// TIA Portal project "TestEssProtoFreia" (V13) (continued)
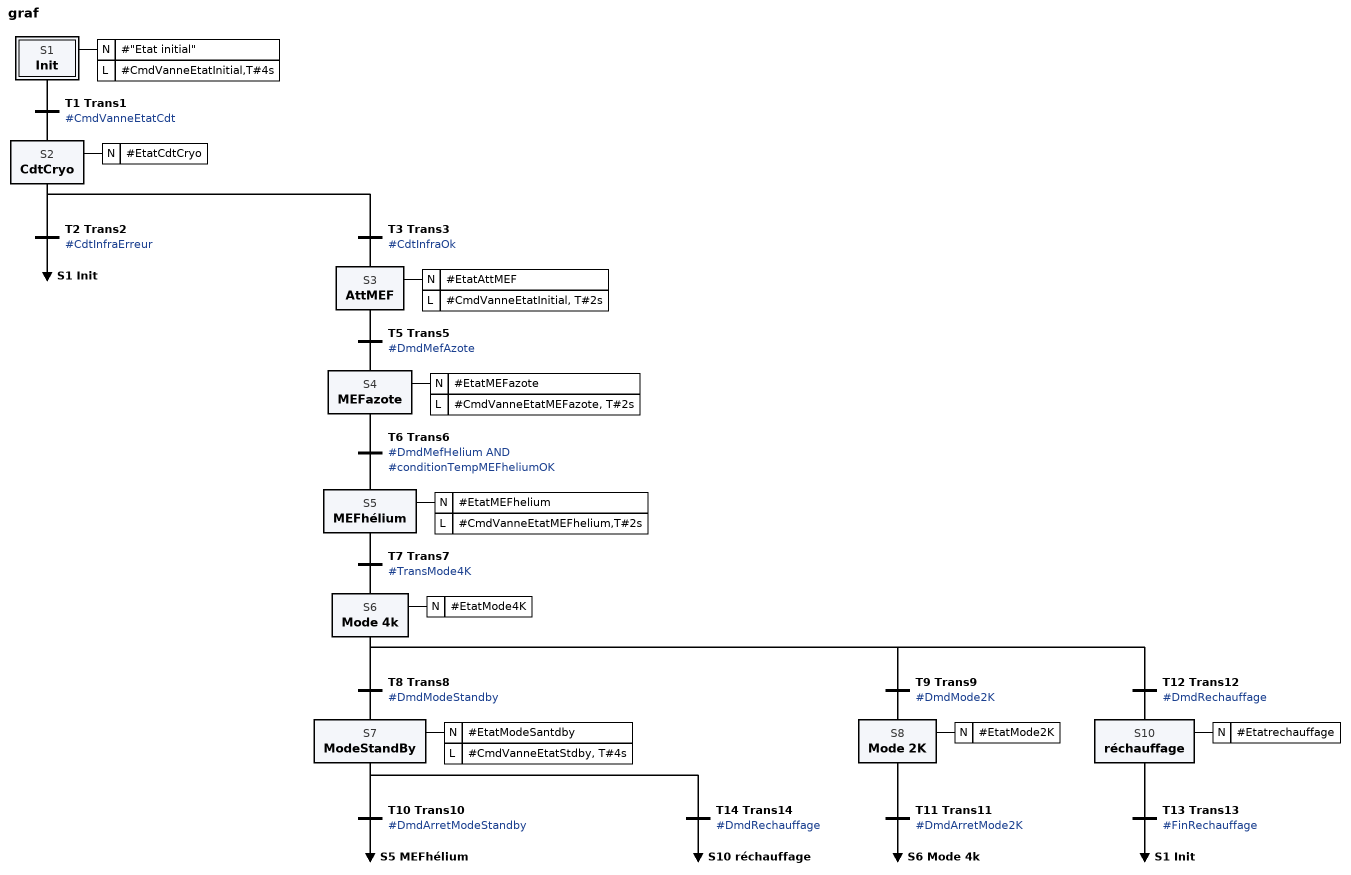
   // sequencer 1
   INITIAL_STEP Init:   // S1
              N    #"Etat initial"
              L    #CmdVanneEtatInitial,T#4s
   END_STEP
   TRANSITION Trans1 FROM Init TO CdtCryo   // T1
      := #CmdVanneEtatCdt;
   END_TRANSITION
   STEP CdtCryo:   // S2
      supervision V := NOT #VanneEnPositionCdt;
      // Version 1: demander manuellement à l automate infra de faire le cdt et confirmer manuellement ( ou pas ) le conditionnement trans3 ( ou trans 2 ) [ajouter boutton cdtinfraok et cdtinfra erreur]
              N    #EtatCdtCryo
   END_STEP
   TRANSITION Trans2 FROM CdtCryo TO Init   // T2, jump
      := #CdtInfraErreur;
   END_TRANSITION
   TRANSITION Trans3 FROM CdtCryo TO AttMEF   // T3
      := #CdtInfraOk;
   END_TRANSITION
   STEP AttMEF:   // S3
      supervision V := NOT #AutorizationMefAzote;
              N    #EtatAttMEF
              L    #CmdVanneEtatInitial, T#2s
   END_STEP
   TRANSITION Trans5 FROM AttMEF TO MEFazote   // T5
      := #DmdMefAzote;
   END_TRANSITION
   STEP MEFazote:   // S4
              N    #EtatMEFazote
              L    #CmdVanneEtatMEFazote, T#2s
   END_STEP
   TRANSITION Trans6 FROM MEFazote TO MEFhélium   // T6
      := #DmdMefHelium AND #conditionTempMEFheliumOK;
   END_TRANSITION
   STEP MEFhélium:   // S5
              N    #EtatMEFhelium
              L    #CmdVanneEtatMEFhelium,T#2s
   END_STEP
   TRANSITION Trans7 FROM MEFhélium TO "Mode 4k"   // T7
      := #TransMode4K;
   END_TRANSITION
   STEP "Mode 4k":   // S6
              N    #EtatMode4K
   END_STEP
   TRANSITION Trans8 FROM "Mode 4k" TO ModeStandBy   // T8
      := #DmdModeStandby;
   END_TRANSITION
   TRANSITION Trans9 FROM "Mode 4k" TO "Mode 2K"   // T9
      := #DmdMode2K;
   END_TRANSITION
   TRANSITION Trans12 FROM "Mode 4k" TO réchauffage   // T12
      := #DmdRechauffage;
   END_TRANSITION
   STEP ModeStandBy:   // S7
              N    #EtatModeSantdby
              L    #CmdVanneEtatStdby, T#4s
   END_STEP
   TRANSITION Trans10 FROM ModeStandBy TO MEFhélium   // T10, jump
      := #DmdArretModeStandby;
   END_TRANSITION
   TRANSITION Trans14 FROM ModeStandBy TO réchauffage   // T14, jump
      := #DmdRechauffage;
   END_TRANSITION
   STEP "Mode 2K":   // S8
              N    #EtatMode2K
   END_STEP
   TRANSITION Trans11 FROM "Mode 2K" TO "Mode 4k"   // T11, jump
      := #DmdArretMode2K;
   END_TRANSITION
   STEP réchauffage:   // S10
              N    #Etatrechauffage
   END_STEP
   TRANSITION Trans13 FROM réchauffage TO Init   // T13, jump
      := #FinRechauffage;
   END_TRANSITION
END_FUNCTION_BLOCK

FUNCTION "commande vanne" : Void   // FC1, LAD
{ S7_Optimized_Access := 'FALSE' }
VERSION : 0.1
   VAR_TEMP   // added for the SCL form of the ladder/FBD networks
      _w1 : Bool;
   END_VAR
BEGIN

REGION Network 1: CV01
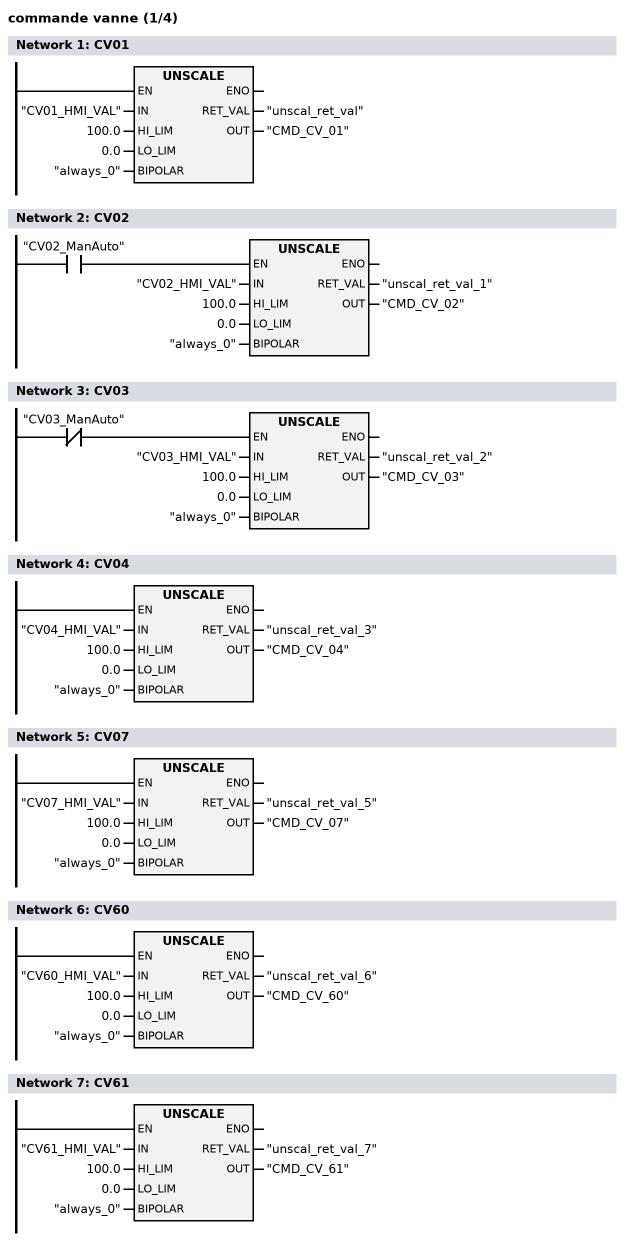
   "unscal_ret_val" := UNSCALE(IN := "CV01_HMI_VAL",
                           HI_LIM := 100.0,
                           LO_LIM := 0.0,
                           BIPOLAR := "always_0",
                           OUT => "CMD_CV_01");
END_REGION

REGION Network 2: CV02
   IF "CV02_ManAuto" THEN
       "unscal_ret_val_1" := UNSCALE(IN := "CV02_HMI_VAL",
                               HI_LIM := 100.0,
                               LO_LIM := 0.0,
                               BIPOLAR := "always_0",
                               OUT => "CMD_CV_02");
   END_IF;
END_REGION

REGION Network 3: CV03
   IF NOT "CV03_ManAuto" THEN
       "unscal_ret_val_2" := UNSCALE(IN := "CV03_HMI_VAL",
                               HI_LIM := 100.0,
                               LO_LIM := 0.0,
                               BIPOLAR := "always_0",
                               OUT => "CMD_CV_03");
   END_IF;
END_REGION

REGION Network 4: CV04
   "unscal_ret_val_3" := UNSCALE(IN := "CV04_HMI_VAL",
                           HI_LIM := 100.0,
                           LO_LIM := 0.0,
                           BIPOLAR := "always_0",
                           OUT => "CMD_CV_04");
END_REGION

REGION Network 5: CV07
   "unscal_ret_val_5" := UNSCALE(IN := "CV07_HMI_VAL",
                           HI_LIM := 100.0,
                           LO_LIM := 0.0,
                           BIPOLAR := "always_0",
                           OUT => "CMD_CV_07");
END_REGION

REGION Network 6: CV60
   "unscal_ret_val_6" := UNSCALE(IN := "CV60_HMI_VAL",
                           HI_LIM := 100.0,
                           LO_LIM := 0.0,
                           BIPOLAR := "always_0",
                           OUT => "CMD_CV_60");
END_REGION

REGION Network 7: CV61
   "unscal_ret_val_7" := UNSCALE(IN := "CV61_HMI_VAL",
                           HI_LIM := 100.0,
                           LO_LIM := 0.0,
                           BIPOLAR := "always_0",
                           OUT => "CMD_CV_61");
END_REGION

REGION Network 8: FT11 (CV11)
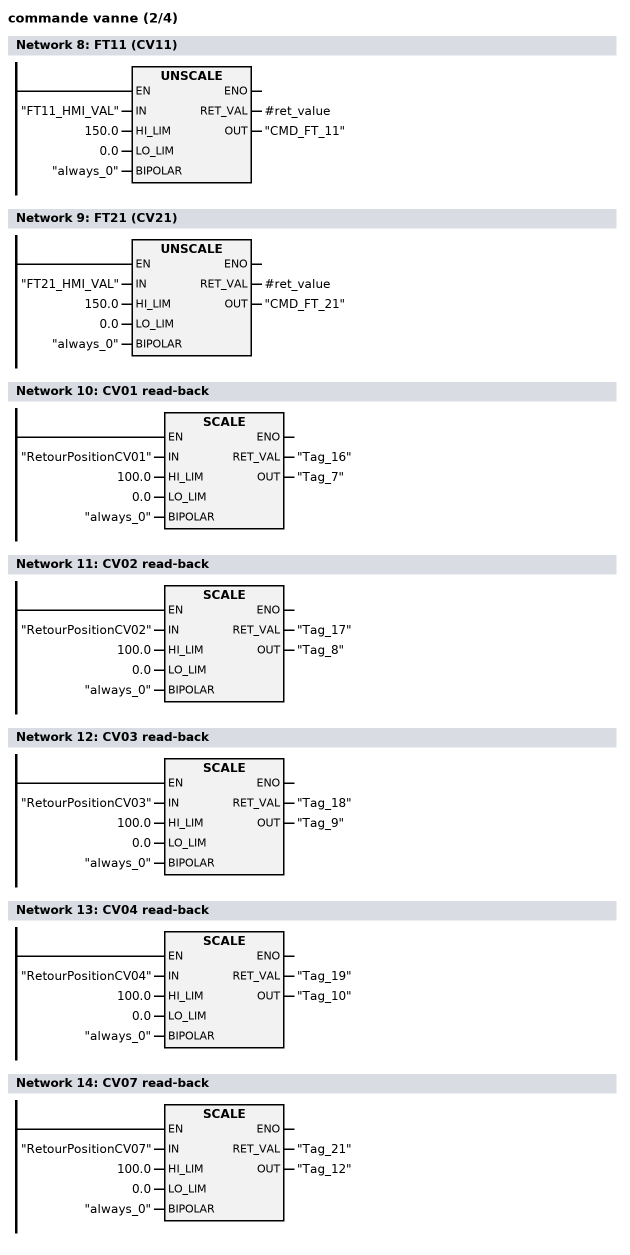
   #ret_value := UNSCALE(IN := "FT11_HMI_VAL",
                         HI_LIM := 150.0,
                         LO_LIM := 0.0,
                         BIPOLAR := "always_0",
                         OUT => "CMD_FT_11");
END_REGION

REGION Network 9: FT21 (CV21)
   #ret_value := UNSCALE(IN := "FT21_HMI_VAL",
                         HI_LIM := 150.0,
                         LO_LIM := 0.0,
                         BIPOLAR := "always_0",
                         OUT => "CMD_FT_21");
END_REGION

REGION Network 10: CV01 read-back
   "Tag_16" := SCALE(IN := "RetourPositionCV01",
                     HI_LIM := 100.0,
                     LO_LIM := 0.0,
                     BIPOLAR := "always_0",
                     OUT => "Tag_7");
END_REGION

REGION Network 11: CV02 read-back
   "Tag_17" := SCALE(IN := "RetourPositionCV02",
                     HI_LIM := 100.0,
                     LO_LIM := 0.0,
                     BIPOLAR := "always_0",
                     OUT => "Tag_8");
END_REGION

REGION Network 12: CV03 read-back
   "Tag_18" := SCALE(IN := "RetourPositionCV03",
                     HI_LIM := 100.0,
                     LO_LIM := 0.0,
                     BIPOLAR := "always_0",
                     OUT => "Tag_9");
END_REGION

REGION Network 13: CV04 read-back
   "Tag_19" := SCALE(IN := "RetourPositionCV04",
                     HI_LIM := 100.0,
                     LO_LIM := 0.0,
                     BIPOLAR := "always_0",
                     OUT => "Tag_10");
END_REGION

REGION Network 14: CV07 read-back
   "Tag_21" := SCALE(IN := "RetourPositionCV07",
                     HI_LIM := 100.0,
                     LO_LIM := 0.0,
                     BIPOLAR := "always_0",
                     OUT => "Tag_12");
END_REGION

REGION Network 15: CV60 read-back
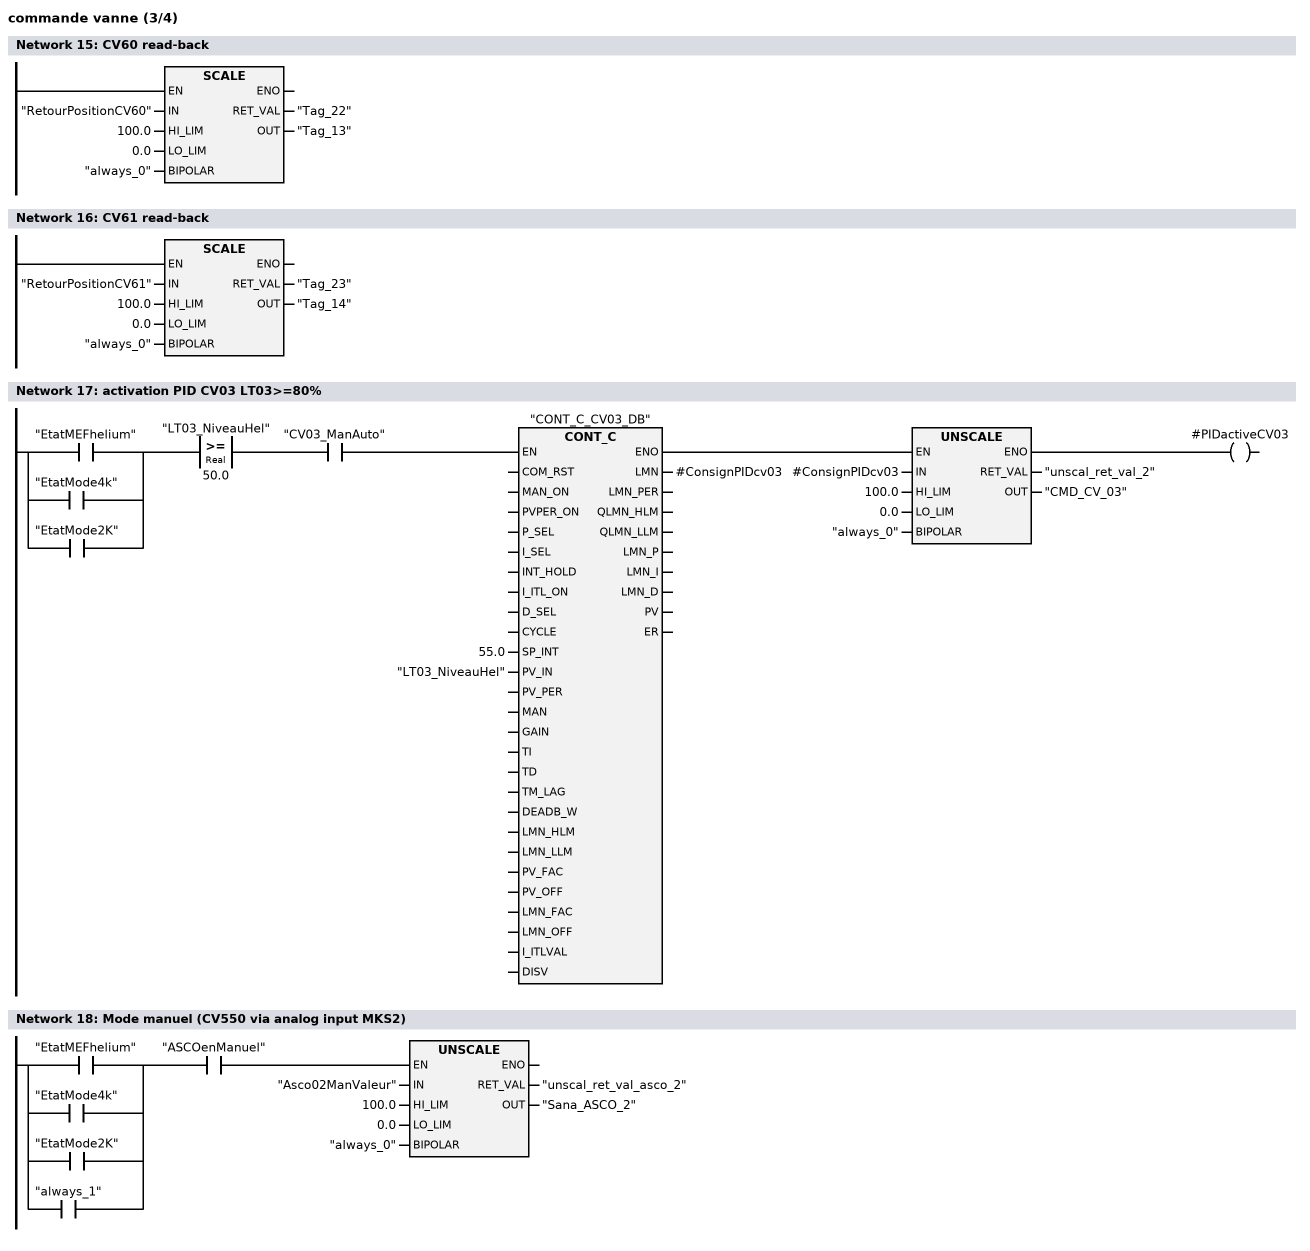
   "Tag_22" := SCALE(IN := "RetourPositionCV60",
                     HI_LIM := 100.0,
                     LO_LIM := 0.0,
                     BIPOLAR := "always_0",
                     OUT => "Tag_13");
END_REGION

REGION Network 16: CV61 read-back
   "Tag_23" := SCALE(IN := "RetourPositionCV61",
                     HI_LIM := 100.0,
                     LO_LIM := 0.0,
                     BIPOLAR := "always_0",
                     OUT => "Tag_14");
END_REGION

REGION Network 17: activation PID CV03 LT03>=80%
   // ENO of a box is taken as its EN; it also drops when the box reports an error
   #_w1 := ("EtatMEFhelium" OR "EtatMode4k" OR "EtatMode2K") AND ("LT03_NiveauHel" >= 50.0) AND "CV03_ManAuto";
   IF #_w1 THEN
       "CONT_C_CV03_DB"(SP_INT := 55.0, PV_IN := "LT03_NiveauHel", LMN => #ConsignPIDcv03);   // CONT_C
       "unscal_ret_val_2" := UNSCALE(IN := #ConsignPIDcv03,
                               HI_LIM := 100.0,
                               LO_LIM := 0.0,
                               BIPOLAR := "always_0",
                               OUT => "CMD_CV_03");
   END_IF;
   #PIDactiveCV03 := #_w1;
END_REGION

REGION Network 18: Mode manuel (CV550 via analog input MKS2)
   IF ("EtatMEFhelium" OR "EtatMode4k" OR "EtatMode2K" OR "always_1") AND "ASCOenManuel" THEN
       "unscal_ret_val_asco_2" := UNSCALE(IN := "Asco02ManValeur",
                               HI_LIM := 100.0,
                               LO_LIM := 0.0,
                               BIPOLAR := "always_0",
                               OUT => "Sana_ASCO_2");
   END_IF;
END_REGION

REGION Network 19: ASCO2 read-back (CV550 read-back via analog output from MKS2)
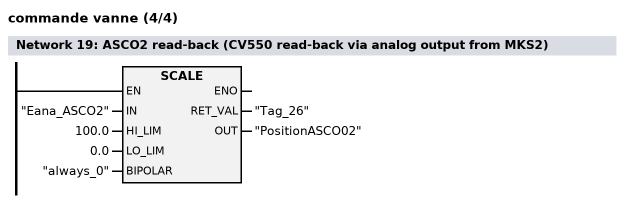
   "Tag_26" := SCALE(IN := "Eana_ASCO2",
                     HI_LIM := 100.0,
                     LO_LIM := 0.0,
                     BIPOLAR := "always_0",
                     OUT => "PositionASCO02");
END_REGION
END_FUNCTION

FUNCTION "NIveau Helium&Pression&vide" : Void   // FC2, STL
{ S7_Optimized_Access := 'FALSE' }
VERSION : 0.1
BEGIN

REGION Network 1: scale niveau helieum LT03
         A     "always_1";
         =     #tmpb;
         BLD   103;
         CALL  "FC10=SCALE"
         ( INPUT       := "Eana_NiveauH_LT03",
           VAL_MAXI    := 74.0,
           VAL_MINI    := 0.0,
           ET_MAX      := 27648,
           ET_MIN      := 0,
           Type_Entree := 0,
           PV_SEUILH   := 100.0,
           PV_SEUILB   := 0.0,
           ACQ         := #tmpb,
           ANIM        := "LT03_TypeDef",
           PV_HIGH     := "LT03_ValMax",
           PV_LOW      := "LT03_ValMin",
           PV          := "LT03_NiveauHel",
           ALM_HIGH    := "LT03_DepHaut",
           ALM_LOW     := "LT03_DepBas",
           ALM_SENSOR  := "LT03_DefSond"
         );
         NOP   0;
END_REGION

REGION Network 2: Copy LT03 to Epics
         L     "LT03_NiveauHel";
         T     "PLC_to_Epics".LT03.Level;
         L     "LT03_TypeDef";
         T     "PLC_to_Epics".LT03.Visu;
         A     "LT03_DefSond";
         =     "PLC_to_Epics".LT03.SensorFlt;
         A     "LT03_DepHaut";
         =     "PLC_to_Epics".LT03.OverRange;
         A     "LT03_DepBas";
         =     "PLC_to_Epics".LT03.UnderRange;
END_REGION

REGION Network 3: scale niveau helieum LT01
         A     "always_1";
         =     #tmpb;
         BLD   103;
         CALL  "FC10=SCALE"
         ( INPUT       := "Eana_NiveauH_LT01",
           VAL_MAXI    := 68.0,
           VAL_MINI    := 0.0,
           ET_MAX      := 27648,
           ET_MIN      := 0,
           Type_Entree := 0,
           PV_SEUILH   := 100.0,
           PV_SEUILB   := 0.0,
           ACQ         := #tmpb,
           ANIM        := "LT01_TypeDef",
           PV_HIGH     := "LT01_ValMax",
           PV_LOW      := "LT01_ValMin",
           PV          := "LT01_NiveauHel",
           ALM_HIGH    := "LT01_DepHaut",
           ALM_LOW     := "LT01_DepBas",
           ALM_SENSOR  := "LT01_DefSond"
         );
         NOP   0;
END_REGION

REGION Network 4: Copy LT01 to Epics
         L     "LT01_NiveauHel";
         T     "PLC_to_Epics".LT01.Level;
         L     "LT01_TypeDef";
         T     "PLC_to_Epics".LT01.Visu;
         A     "LT01_DefSond";
         =     "PLC_to_Epics".LT01.SensorFlt;
         A     "LT01_DepHaut";
         =     "PLC_to_Epics".LT01.OverRange;
         A     "LT01_DepBas";
         =     "PLC_to_Epics".LT01.UnderRange;
END_REGION

REGION Network 5: scale niveau helieum LT02
         A     "always_1";
         =     #tmpb;
         BLD   103;
         CALL  "FC10=SCALE"
         ( INPUT       := "Eana_NiveauH_LT02",
           VAL_MAXI    := 68.0,
           VAL_MINI    := 0.0,
           ET_MAX      := 27648,
           ET_MIN      := 0,
           Type_Entree := 0,
           PV_SEUILH   := 100.0,
           PV_SEUILB   := 0.0,
           ACQ         := #tmpb,
           ANIM        := "LT02_TypeDef",
           PV_HIGH     := "LT02_ValMax",
           PV_LOW      := "LT02_ValMin",
           PV          := "LT02_NiveauHel",
           ALM_HIGH    := "LT02_DepHaut",
           ALM_LOW     := "LT02_DepBas",
           ALM_SENSOR  := "LT02_DefSond"
         );
         NOP   0;
END_REGION

REGION Network 6: Copy LT02 to Epics
         L     "LT02_NiveauHel";
         T     "PLC_to_Epics".LT02.Level;
         L     "LT02_TypeDef";
         T     "PLC_to_Epics".LT02.Visu;
         A     "LT02_DefSond";
         =     "PLC_to_Epics".LT02.SensorFlt;
         A     "LT02_DepHaut";
         =     "PLC_to_Epics".LT02.OverRange;
         A     "LT02_DepBas";
         =     "PLC_to_Epics".LT02.UnderRange;
END_REGION

REGION Network 7: Set an interlock signal for RF slow interlock
         AN    "LT01_DefSond";
         AN    "LT01_DepHaut";
         AN    "LT01_DepBas";
         A(;
         L     "LT01_NiveauHel";
         L     50.0;
         >R;
         );
         =     "CM_CryoOK";
END_REGION

REGION Network 8: scale pression PT60 ecran thermique
         A     "always_0";
         =     #tmpb;
         BLD   103;
         CALL  SCALE
         ( IN      := "Eana_PressionPT60",
           HI_LIM  := 2660.0,
           LO_LIM  := 0.0,
           BIPOLAR := #tmpb,
           RET_VAL := "ScaleErreurPT60",
           OUT     := "Pression".PressionPT60_Val
         );
         NOP   0;
END_REGION

REGION Network 9: Copy PT60 to Epics
         L     "Pression".PressionPT60_Val;
         T     "PLC_to_Epics".PT60;
END_REGION

REGION Network 10: scale pression PT01
         A     "always_0";
         =     #tmpb;
         BLD   103;
         CALL  SCALE
         ( IN      := "Eana_PressionPT01",
           HI_LIM  := 2660.0,
           LO_LIM  := 0.0,
           BIPOLAR := #tmpb,
           RET_VAL := "ScaleErreurPT01",
           OUT     := "Pression".PressionPT01_Val
         );
         NOP   0;
END_REGION

REGION Network 11: Copy PT01 to Epics
         L     "Pression".PressionPT01_Val;
         T     "PLC_to_Epics".PT01;
END_REGION

REGION Network 12: scale pression diff
         A     "always_1";
         =     #tmpb;
         BLD   103;
         CALL  SCALE
         ( IN      := "Eana_PressionDiff",
           HI_LIM  := 1.33322,
           LO_LIM  := -1.33322,
           BIPOLAR := #tmpb,
           RET_VAL := "ScaleErreurPressionDiff",
           OUT     := "Pression".PressionDiff
         );
         NOP   0;
END_REGION

REGION Network 13: Copy PT04 to Epics
         L     "Pression".PressionDiff;
         T     "PLC_to_Epics".PT04;
END_REGION

REGION Network 14: sclae vide VB PT73
         A     "always_0";
         =     #tmpb;
         BLD   103;
         CALL  SCALE
         ( IN      := "Eana_VidePT73",
           HI_LIM  := 10.0,
           LO_LIM  := 0.0,
           BIPOLAR := #tmpb,
           RET_VAL := "ScaleErreurVidePT73",
           OUT     := "VidePT73Tension"
         );
         NOP   0;
END_REGION

REGION Network 15: Tension / Pression Vide PT73
         CALL  "CALCUL VIDE"
         ( VOLT     := "VidePT73Tension",
           PRESSION := "Pression".PressionVidePT73
         );
         NOP   0;
END_REGION

REGION Network 16: Copy PT73 to Epics
         L     "Pression".PressionVidePT73;
         T     "PLC_to_Epics".PT73;
END_REGION

REGION Network 17: scale vide CM PT71
         A     "always_0";
         =     #tmpb;
         BLD   103;
         CALL  SCALE
         ( IN      := "Eana_VidePT71",
           HI_LIM  := 10.0,
           LO_LIM  := 0.0,
           BIPOLAR := #tmpb,
           RET_VAL := "ScaleErreurVidePT71",
           OUT     := "VidePT71Tension"
         );
         NOP   0;
END_REGION

REGION Network 18: Tension / Pression Vide PT71
         CALL  "CALCUL VIDE"
         ( VOLT     := "VidePT71Tension",
           PRESSION := "Pression".PressionVidePT71
         );
         NOP   0;
END_REGION

REGION Network 19: Copy PT71 to Epics
         L     "Pression".PressionVidePT71;
         T     "PLC_to_Epics".PT71;
END_REGION

REGION Network 20: Scale vide PT75
         A     "always_0";
         =     #tmpb;
         BLD   103;
         CALL  SCALE
         ( IN      := "Eana_VidePT75",
           HI_LIM  := 10.0,
           LO_LIM  := 0.0,
           BIPOLAR := #tmpb,
           RET_VAL := "Tag_50",
           OUT     := "Tag_48"
         );
         NOP   0;
END_REGION

REGION Network 21: Calcul pression PT75
         CALL  "CALCUL VIDE"
         ( VOLT     := "Tag_48",
           PRESSION := "Pression".PressionVidePT75
         );
         NOP   0;
END_REGION

REGION Network 22: Copy PT75 to Epics
         L     "Pression".PressionVidePT75;
         T     "PLC_to_Epics".PT75;
END_REGION

REGION Network 23: scale PT77
         A     "always_0";
         =     #tmpb;
         BLD   103;
         CALL  SCALE
         ( IN      := "Eana_VidePT77",
           HI_LIM  := 10.0,
           LO_LIM  := 0.0,
           BIPOLAR := #tmpb,
           RET_VAL := "Tag_51",
           OUT     := "Tag_52"
         );
         NOP   0;
END_REGION

REGION Network 24: Calcul Pression PT77
         CALL  "CALCUL VIDE"
         ( VOLT     := "Tag_52",
           PRESSION := "Pression".PressionVidePT77
         );
         NOP   0;
END_REGION

REGION Network 25: Copy PT77 to Epics
         L     "Pression".PressionVidePT77;
         T     "PLC_to_Epics".PT77;
END_REGION

REGION Network 26: FT11 - scale and copy to Epics
         A     "always_1";
         =     #tmpb;
         BLD   103;
         CALL  "FC10=SCALE"
         ( INPUT       := "FT11",
           VAL_MAXI    := 150.0,
           VAL_MINI    := -0.542534,
           ET_MAX      := 27648,
           ET_MIN      := -100,
           Type_Entree := 0,
           PV_SEUILH   := 150.0,
           PV_SEUILB   := -0.5,
           ACQ         := #tmpb,
           ANIM        := "PLC_to_Epics".FT11.Visu,
           PV_HIGH     := #tmpr,
           PV_LOW      := #tmpr,
           PV          := "PLC_to_Epics".FT11.Level,
           ALM_HIGH    := "PLC_to_Epics".FT11.OverRange,
           ALM_LOW     := "PLC_to_Epics".FT11.UnderRange,
           ALM_SENSOR  := "PLC_to_Epics".FT11.SensorFlt
         );

         NOP   0;
END_REGION

REGION Network 27: FT21 - scale and copy to Epics
         A     "always_1";
         =     #tmpb;
         BLD   103;
         CALL  "FC10=SCALE"
         ( INPUT       := "FT21",
           VAL_MAXI    := 150.0,
           VAL_MINI    := -0.542534,
           ET_MAX      := 27648,
           ET_MIN      := -100,
           Type_Entree := 0,
           PV_SEUILH   := 150.0,
           PV_SEUILB   := -0.5,
           ACQ         := #tmpb,
           ANIM        := "PLC_to_Epics".FT21.Visu,
           PV_HIGH     := #tmpr,
           PV_LOW      := #tmpr,
           PV          := "PLC_to_Epics".FT21.Level,
           ALM_HIGH    := "PLC_to_Epics".FT21.OverRange,
           ALM_LOW     := "PLC_to_Epics".FT21.UnderRange,
           ALM_SENSOR  := "PLC_to_Epics".FT21.SensorFlt
         );
         NOP   0;
END_REGION

REGION Network 28: TT110 - scale and copy to Epics
         A     "always_1";
         =     #tmpb;
         BLD   103;
         CALL  "FC10=SCALE"
         ( INPUT       := "TT110",
           VAL_MAXI    := 373.15,
           VAL_MINI    := 93.15,
           ET_MAX      := 27648,
           ET_MIN      := 0,
           Type_Entree := 0,
           PV_SEUILH   := 373.15,
           PV_SEUILB   := 93.15,
           ACQ         := #tmpb,
           ANIM        := "PLC_to_Epics".TT110.Visu,
           PV_HIGH     := #tmpr,
           PV_LOW      := #tmpr,
           PV          := "PLC_to_Epics".TT110.Level,
           ALM_HIGH    := "PLC_to_Epics".TT110.OverRange,
           ALM_LOW     := "PLC_to_Epics".TT110.UnderRange,
           ALM_SENSOR  := "PLC_to_Epics".TT110.SensorFlt
         );
         NOP   0;
END_REGION

REGION Network 29: TT210 - scale and copy to Epics
         A     "always_1";
         =     #tmpb;
         BLD   103;
         CALL  "FC10=SCALE"
         ( INPUT       := "TT210",
           VAL_MAXI    := 373.15,
           VAL_MINI    := 93.15,
           ET_MAX      := 27648,
           ET_MIN      := 0,
           Type_Entree := 0,
           PV_SEUILH   := 373.15,
           PV_SEUILB   := 93.15,
           ACQ         := #tmpb,
           ANIM        := "PLC_to_Epics".TT210.Visu,
           PV_HIGH     := #tmpr,
           PV_LOW      := #tmpr,
           PV          := "PLC_to_Epics".TT210.Level,
           ALM_HIGH    := "PLC_to_Epics".TT210.OverRange,
           ALM_LOW     := "PLC_to_Epics".TT210.UnderRange,
           ALM_SENSOR  := "PLC_to_Epics".TT210.SensorFlt
         );
         NOP   0;
END_REGION

REGION Network 30: Copy PT02_direct to Epics
         L     "Pression".PT02_direct;
         T     "PLC_to_Epics".PT02_direct;
END_REGION
END_FUNCTION

FUNCTION "ACQ_CABTF" : Void   // FC3, STL
{ S7_Optimized_Access := 'FALSE' }
VERSION : 0.1
BEGIN

REGION Network 1: Copy data from CATBF1 to Epics
         CALL  BLKMOV
         ( SRCBLK  := P#I518.0 WORD 16,
           RET_VAL := #Fault_de_la_Copie,
           DSTBLK  := "PLC_to_Epics".CABTF1.board1
         );
         CALL  BLKMOV
         ( SRCBLK  := P#I582.0 WORD 16,
           RET_VAL := #Fault_de_la_Copie,
           DSTBLK  := "PLC_to_Epics".CABTF1.board2
         );
         CALL  BLKMOV
         ( SRCBLK  := P#I646.0 WORD 4,
           RET_VAL := #Fault_de_la_Copie,
           DSTBLK  := "PLC_to_Epics".CABTF1.stat
         );
END_REGION

REGION Network 2: Copy data from CATBF2 to Epics
         CALL  BLKMOV
         ( SRCBLK  := P#I716.0 WORD 16,
           RET_VAL := #Fault_de_la_Copie,
           DSTBLK  := "PLC_to_Epics".CABTF2.board1
         );
         CALL  BLKMOV
         ( SRCBLK  := P#I780.0 WORD 16,
           RET_VAL := #Fault_de_la_Copie,
           DSTBLK  := "PLC_to_Epics".CABTF2.board2
         );
         CALL  BLKMOV
         ( SRCBLK  := P#I472.0 WORD 4,
           RET_VAL := #Fault_de_la_Copie,
           DSTBLK  := "PLC_to_Epics".CABTF2.stat
         );
END_REGION

REGION Network 3: Copy data from CATBF3 to Epics
         CALL  BLKMOV
         ( SRCBLK  := P#I336.0 WORD 32,
           RET_VAL := #Fault_de_la_Copie,
           DSTBLK  := "PLC_to_Epics".CABTF3
         );
         CALL  BLKMOV
         ( SRCBLK  := P#I400.0 WORD 16,
           RET_VAL := #Fault_de_la_Copie,
           DSTBLK  := "PLC_to_Epics".CABTF3.board2
         );
         CALL  BLKMOV
         ( SRCBLK  := P#I464.0 WORD 4,
           RET_VAL := #Fault_de_la_Copie,
           DSTBLK  := "PLC_to_Epics".CABTF3.stat
         );
END_REGION

REGION Network 4: TT77
         A     "always_1";
         =     #tmpb;
         BLD   103;
         CALL  "FC10=SCALE"
         ( INPUT       := "Eana_TT77_ohm",
           VAL_MAXI    := 150.0,
           VAL_MINI    := 0.0,
           ET_MAX      := 27648,
           ET_MIN      := 0,
           Type_Entree := 0,
           PV_SEUILH   := 400.0,
           PV_SEUILB   := 0.0,
           ACQ         := #tmpb,
           ANIM        := "tt77typedef",
           PV_HIGH     := "tt77max",
           PV_LOW      := "tt77min",
           PV          := "ReceivePT100"."TT77_(R)",
           ALM_HIGH    := "tt77h",
           ALM_LOW     := "tt77l",
           ALM_SENSOR  := "tt77alm"
         );
         NOP   0;
END_REGION

REGION Network 5: TT77 - convert R -> T
         CALL  "CONVERSION R/T"
         ( "RESISTANCE _OHMS" := "ReceivePT100"."TT77_(R)",
           TEMPERATURE_KELVIN := "ReceivePT100"."TT77_(K)"
         );
         NOP   0;
END_REGION

REGION Network 6: Copy TT77 to Epics
         L     "ReceivePT100"."TT77_(K)";
         T     "PLC_to_Epics".TT77.Level;
         L     "tt77typedef";
         T     "PLC_to_Epics".TT77.Visu;
         A     "tt77alm";
         =     "PLC_to_Epics".TT77.SensorFlt;
         A     "tt77h";
         =     "PLC_to_Epics".TT77.OverRange;
         A     "tt77l";
         =     "PLC_to_Epics".TT77.UnderRange;
END_REGION

REGION Network 7: TT120 - scale and fill epics buffer
         A     "always_1";
         =     #tmpb;
         BLD   103;
         CALL  "FC10=SCALE"
         ( INPUT       := "TT120",
           VAL_MAXI    := 150.0,
           VAL_MINI    := 0.0,
           ET_MAX      := 27648,
           ET_MIN      := 0,
           Type_Entree := 0,
           PV_SEUILH   := 400.0,
           PV_SEUILB   := 0.0,
           ACQ         := #tmpb,
           ANIM        := "PLC_to_Epics".TT120.Visu,
           PV_HIGH     := #tmpr,
           PV_LOW      := #tmpr,
           PV          := #resistance,
           ALM_HIGH    := "PLC_to_Epics".TT120.OverRange,
           ALM_LOW     := "PLC_to_Epics".TT120.UnderRange,
           ALM_SENSOR  := "PLC_to_Epics".TT120.SensorFlt
         );
         NOP   0;
END_REGION

REGION Network 8: TT120 - convert R -> T
         CALL  "CONVERSION R/T"
         ( "RESISTANCE _OHMS" := #resistance,
           TEMPERATURE_KELVIN := "PLC_to_Epics".TT120.Level
         );
         NOP   0;
END_REGION

REGION Network 9: TT220 - scale and fill epics buffer
         A     "always_1";
         =     #tmpb;
         BLD   103;
         CALL  "FC10=SCALE"
         ( INPUT       := "TT220",
           VAL_MAXI    := 150.0,
           VAL_MINI    := 0.0,
           ET_MAX      := 27648,
           ET_MIN      := 0,
           Type_Entree := 0,
           PV_SEUILH   := 400.0,
           PV_SEUILB   := 0.0,
           ACQ         := #tmpb,
           ANIM        := "PLC_to_Epics".TT220.Visu,
           PV_HIGH     := #tmpr,
           PV_LOW      := #tmpr,
           PV          := #resistance,
           ALM_HIGH    := "PLC_to_Epics".TT220.OverRange,
           ALM_LOW     := "PLC_to_Epics".TT220.UnderRange,
           ALM_SENSOR  := "PLC_to_Epics".TT220.SensorFlt
         );
         NOP   0;
END_REGION

REGION Network 10: TT220 - convert R -> T
         CALL  "CONVERSION R/T"
         ( "RESISTANCE _OHMS" := #resistance,
           TEMPERATURE_KELVIN := "PLC_to_Epics".TT220.Level
         );
         NOP   0;
END_REGION
END_FUNCTION

FUNCTION "CALCUL VIDE" : Void   // FC4, SCL
{ S7_Optimized_Access := 'FALSE' }
VERSION : 0.1
BEGIN

   #PRESSION := 10 ** ((1.667*#VOLT) - 11.33);
END_FUNCTION

FUNCTION "PID ASCO" : Void   // FC5, LAD
{ S7_Optimized_Access := 'FALSE' }
VERSION : 0.1
   VAR_TEMP   // added for the SCL form of the ladder/FBD networks
      _w1 : Bool;
   END_VAR
BEGIN

REGION Network 1: PID ASCO 2
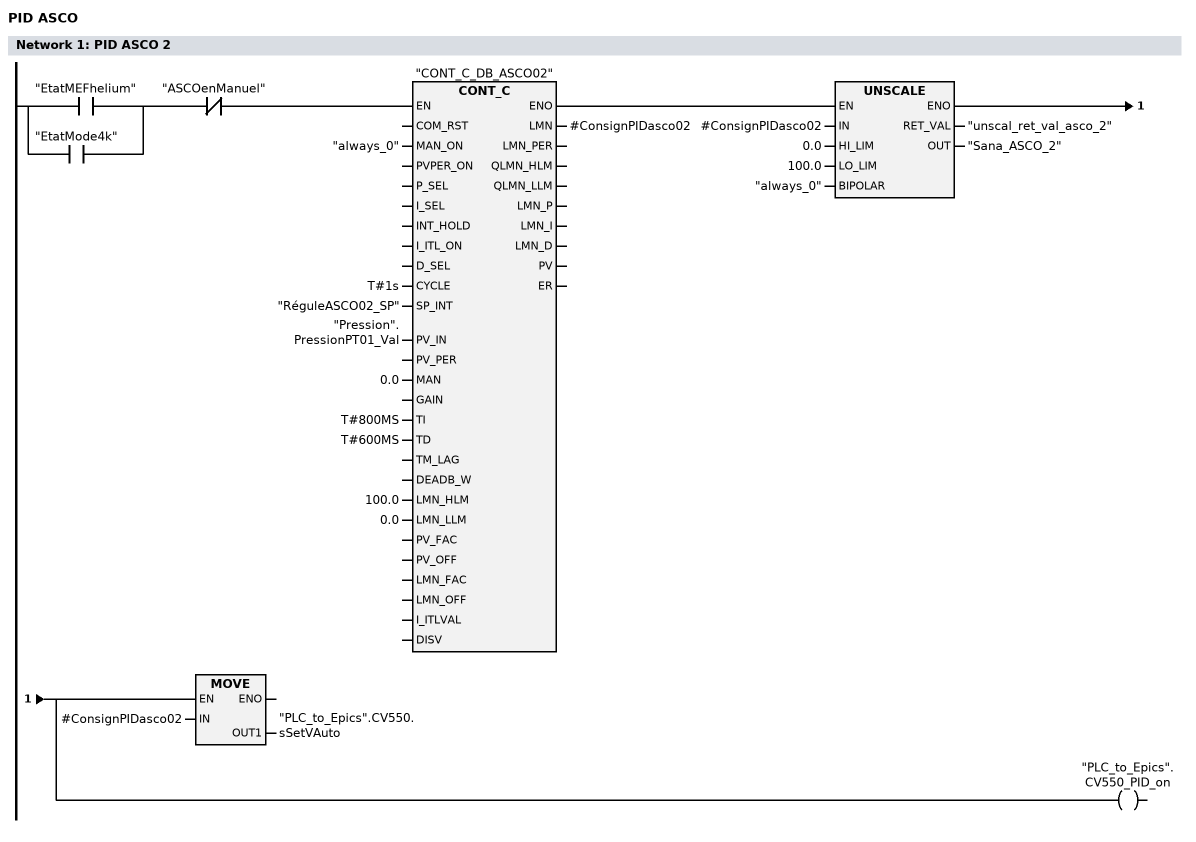
   // ENO of a box is taken as its EN; it also drops when the box reports an error
   #_w1 := ("EtatMEFhelium" OR "EtatMode4k") AND NOT "ASCOenManuel";
   IF #_w1 THEN
       "CONT_C_DB_ASCO02"(MAN_ON := "always_0",   // CONT_C
                          CYCLE := T#1s,
                          SP_INT := "RéguleASCO02_SP",
                          PV_IN := "Pression".PressionPT01_Val,
                          MAN := 0.0,
                          TI := T#800MS,
                          TD := T#600MS,
                          LMN_HLM := 100.0,
                          LMN_LLM := 0.0,
                          LMN => #ConsignPIDasco02);
       "unscal_ret_val_asco_2" := UNSCALE(IN := #ConsignPIDasco02,
                               HI_LIM := 0.0,
                               LO_LIM := 100.0,
                               BIPOLAR := "always_0",
                               OUT => "Sana_ASCO_2");
       "PLC_to_Epics".CV550.sSetVAuto := #ConsignPIDasco02;
   END_IF;
   "PLC_to_Epics".CV550_PID_on := #_w1;
END_REGION
END_FUNCTION

FUNCTION "FC10=SCALE" : Void   // FC10, FBD
TITLE = SCALE
{ S7_Optimized_Access := 'FALSE' }
VERSION : 0.1
BEGIN

REGION Network 1 (STL): input type select
         L     #Type_Entree;
         JL    LSTX;
         JU    C1;  // Valeur 0 : Tension ou courant
         JU    C2;  // Valeur 1 : PT100 en °C
         JU    C3;  // Valeur 2 : PT100 en K
   LSTX: JU    End;
END_REGION

REGION Network 2 (STL): Input type : 4-20mA, 0/10V
   // Input type  : 4-20mA, 0/10V
   // 
   // (Acquisition - Etendue mesure mini)*(Echelle max - min) + Echelle mini = mesure 
   // convertie
   // 
   // Etendue mesure maxi - mini
   C1:   L     #INPUT;
         ITD;
         DTR;
         L     #ET_MIN;
         ITD;
         DTR;
         -R;
         T     #INTER_1;  //Acquisition - etendue de mesure mini

         L     #VAL_MAXI;
         L     #VAL_MINI;
         -R;
         T     #INTER_2;  //ECHELLE MAXI - MINI